      Visibility <- "DB939_Tool_alloc_HMI_Limit_allocation_list"
   Button "Button_96" at 118,470 size 306x41; TextOff 'Text'
      on Press: SetTag("DB939_Tool_alloc_HMI_Selected_prog", 9)
      Visibility <- "DB939_Tool_alloc_HMI_Limit_allocation_list"
   Button "Button_97" at 118,510 size 306x41; TextOff 'Text'
      on Press: SetTag("DB939_Tool_alloc_HMI_Selected_prog", 10)
      Visibility <- "DB939_Tool_alloc_HMI_Limit_allocation_list"
   Button "Button_98" at 118,550 size 306x41; TextOff 'Text'
      on Press: SetTag("DB939_Tool_alloc_HMI_Selected_prog", 11)
      Visibility <- "DB939_Tool_alloc_HMI_Limit_allocation_list"
   Button "Button_99" at 118,590 size 306x41; TextOff 'Text'
      on Press: SetTag("DB939_Tool_alloc_HMI_Selected_prog", 12)
      Visibility <- "DB939_Tool_alloc_HMI_Limit_allocation_list"
   Button "Button_100" at 118,630 size 306x41; TextOff 'Text'
      on Press: SetTag("DB939_Tool_alloc_HMI_Selected_prog", 13)
      Visibility <- "DB939_Tool_alloc_HMI_Limit_allocation_list"
   Button "Button_101" at 118,670 size 306x41; TextOff 'Text'
      on Press: SetTag("DB939_Tool_alloc_HMI_Selected_prog", 14)
      Visibility <- "DB939_Tool_alloc_HMI_Limit_allocation_list"
   Button "Button_102" at 118,710 size 306x41; TextOff 'Text'
      on Press: SetTag("DB939_Tool_alloc_HMI_Selected_prog", 15)
      Visibility <- "DB939_Tool_alloc_HMI_Limit_allocation_list"
   Button "Button_103" at 491,149 size 306x41; TextOff 'Text'
      on Press: SetTag("DB939_Tool_alloc_HMI_Selected_prog", 16)
      Visibility <- "DB939_Tool_alloc_HMI_Limit_allocation_list"
   Button "Button_104" at 491,189 size 306x41; TextOff 'Text'
      on Press: SetTag("DB939_Tool_alloc_HMI_Selected_prog", 17)
      Visibility <- "DB939_Tool_alloc_HMI_Limit_allocation_list"
   Button "Button_105" at 491,229 size 306x41; TextOff 'Text'
      on Press: SetTag("DB939_Tool_alloc_HMI_Selected_prog", 18)
      Visibility <- "DB939_Tool_alloc_HMI_Limit_allocation_list"
   Button "Button_106" at 491,269 size 306x41; TextOff 'Text'
      on Press: SetTag("DB939_Tool_alloc_HMI_Selected_prog", 19)
      Visibility <- "DB939_Tool_alloc_HMI_Limit_allocation_list"
   Button "Button_107" at 491,309 size 306x41; TextOff 'Text'
      on Press: SetTag("DB939_Tool_alloc_HMI_Selected_prog", 20)
      Visibility <- "DB939_Tool_alloc_HMI_Limit_allocation_list"
   Button "Button_108" at 491,349 size 306x41; TextOff 'Text'
      on Press: SetTag("DB939_Tool_alloc_HMI_Selected_prog", 21)
      Visibility <- "DB939_Tool_alloc_HMI_Limit_allocation_list"
   Button "Button_109" at 491,389 size 306x41; TextOff 'Text'
      on Press: SetTag("DB939_Tool_alloc_HMI_Selected_prog", 22)
      Visibility <- "DB939_Tool_alloc_HMI_Limit_allocation_list"
   Button "Button_110" at 491,429 size 306x41; TextOff 'Text'
      on Press: SetTag("DB939_Tool_alloc_HMI_Selected_prog", 23)
      Visibility <- "DB939_Tool_alloc_HMI_Limit_allocation_list"
   Button "Button_111" at 491,469 size 306x41; TextOff 'Text'
      on Press: SetTag("DB939_Tool_alloc_HMI_Selected_prog", 24)
      Visibility <- "DB939_Tool_alloc_HMI_Limit_allocation_list"
   Button "Button_112" at 491,509 size 306x41; TextOff 'Text'
      on Press: SetTag("DB939_Tool_alloc_HMI_Selected_prog", 25)
      Visibility <- "DB939_Tool_alloc_HMI_Limit_allocation_list"
   Button "Button_113" at 491,549 size 306x41; TextOff 'Text'
      on Press: SetTag("DB939_Tool_alloc_HMI_Selected_prog", 26)
      Visibility <- "DB939_Tool_alloc_HMI_Limit_allocation_list"
   Button "Button_114" at 491,589 size 306x41; TextOff 'Text'
      on Press: SetTag("DB939_Tool_alloc_HMI_Selected_prog", 27)
      Visibility <- "DB939_Tool_alloc_HMI_Limit_allocation_list"
   Button "Button_115" at 491,629 size 306x41; TextOff 'Text'
      on Press: SetTag("DB939_Tool_alloc_HMI_Selected_prog", 28)
      Visibility <- "DB939_Tool_alloc_HMI_Limit_allocation_list"
   Button "Button_116" at 491,669 size 306x41; TextOff 'Text'
      on Press: SetTag("DB939_Tool_alloc_HMI_Selected_prog", 29)
      Visibility <- "DB939_Tool_alloc_HMI_Limit_allocation_list"
   Button "Button_117" at 491,709 size 306x41; TextOff 'Text'
      on Press: SetTag("DB939_Tool_alloc_HMI_Selected_prog", 30)
      Visibility <- "DB939_Tool_alloc_HMI_Limit_allocation_list"

screen "0013_Archive Alarm" 1280x800, template "Navigation"
   on GenerateScreen: SetTag("CopyLogControl", 0)
   on ClearScreen: SetTag("NavScreenChange", 0); SetTag("CopyLogControl", 0)
   AlarmView "Alarm Archived Fault" at 108,175 size 1058x498; AlarmLog "Archivanzeige"
      Visibility <- "Archived Alarm Control"
   Button "b_System" at 799,713 size 60x60; TextOff 'System'; PictureOff "system messages"; TextList "ico"; PictureList "ico_System_message"
      Appearance <- "Archived Alarm Control"
      on Click: SetTag("Archived Alarm Control", 3)
      ProcessValue <- "Archived Alarm Control"
   Button "b_Foaming" at 891,712 size 60x60; TextOff 'Foaming'; PictureList "ico_Foaming"
      Appearance <- "Archived Alarm Control"
      on Click: SetTag("Archived Alarm Control", 2)
      ProcessValue <- "Archived Alarm Control"
   Button "b_FaultFoam" at 984,712 size 60x60; TextOff 'Fault/Foam'; PictureList "ico_ActualFault_Foaming"
      Appearance <- "Archived Alarm Control"
      on Click: SetTag("Archived Alarm Control", 1)
      ProcessValue <- "Archived Alarm Control"
   Button "b_Fault" at 1077,712 size 60x60; TextOff 'Fault'; PictureList "ico_Actual_Fault"
      Appearance <- "Archived Alarm Control"
      on Click: SetTag("Archived Alarm Control", 0)
      ProcessValue <- "Archived Alarm Control"
   Button "Button_3" at 326,104 size 451x32; TextOff 'Actual Fault / foaming data'; TextList "Archived_Screen_Name_List"
      ProcessValue <- "Archived Alarm Control"
   Button "b_USB" at 705,712 size 60x60; TextOff 'Export USB'; PictureOff "USB_1"
      on Click: function_e9be9208(1, "Archivanzeige", '\Storage Card USB\', 0)
   Button "b_Fault_1" at 1077,712 size 60x60; TextOff 'Fault'
      on Click: SetTag("Archived Alarm Control", 0)
      Appearance <- "Archived Alarm Control"
   Button "b_Foaming_1" at 891,712 size 60x60; TextOff 'Foaming'
      on Click: SetTag("Archived Alarm Control", 2)
      Appearance <- "Archived Alarm Control"
   Button "b_FaultFoam_1" at 984,712 size 60x60; TextOff 'Fault/Foam'
      on Click: SetTag("Archived Alarm Control", 1)
      Appearance <- "Archived Alarm Control"
   Button "b_System_1" at 799,713 size 60x60; TextOff 'System'; PictureOff "system messages"
      on Click: SetTag("Archived Alarm Control", 3)
      Appearance <- "Archived Alarm Control"
   Button "b_ShifProto_ShotCounter_1" at 208,713 size 60x60; TextOff 'Shot Counter'; PictureList "ico_ShiftProtocol"
      ProcessValue <- "Recipe_Appearance_Control"
      Appearance <- "Recipe_Appearance_Control"
   Button "b_Shiftproto_shiftproto" at 208,713 size 60x60; TextOff 'Shift proto'
      on Click: ActivateScreen("0112_Shift protocol", 0); SetTag("Recipe_Appearance_Control", 2)
      Appearance <- "Recipe_Appearance_Control"
   Button "b_SC" at 478,713 size 60x60; TextOff 'Shot Counter'; PictureList "ico_ShotCounter"
      on Press: ActivateScreen("0891_Shotcounter MixingHead", 0); SetTag("Recipe_Appearance_Control", 5)
      Appearance <- "Recipe_Appearance_Control"
      ProcessValue <- "Recipe_Appearance_Control"
   Button "b_SC_1" at 478,713 size 60x60; TextOff 'Shot Counter'
      on Click: ActivateScreen("0891_Shotcounter MixingHead", 0); SetTag("Recipe_Appearance_Control", 5)
      Appearance <- "Recipe_Appearance_Control"
   Button "b_Shift_Plan" at 118,713 size 60x60; TextOff 'Shift Plan'; PictureList "ico_ShiftPlan"
      on Press: ActivateScreen("0113_SettingShiftPlan", 0); SetTag("Recipe_Appearance_Control", 1)
      Appearance <- "Recipe_Appearance_Control"
      ProcessValue <- "Recipe_Appearance_Control"
   Button "b_Shift_Plan_1" at 118,713 size 60x60; TextOff 'Shift Plan'
      on Click: "SettingShiftPlan"(); ActivateScreen("0113_SettingShiftPlan", 0); SetTag("Recipe_Appearance_Control", 1)
      Appearance <- "Recipe_Appearance_Control"
   Button "b_LS_Lastshot" at 298,713 size 60x60; TextOff 'Last Shot'; PictureList "ico_LastShot"
      on Press: ActivateScreen("0036_Last Shot", 0); SetTag("Recipe_Appearance_Control", 3)
      Appearance <- "Recipe_Appearance_Control"
      ProcessValue <- "Recipe_Appearance_Control"
   Button "b_LS_Lastshot_1" at 298,713 size 60x60; TextOff 'Last Shot'
      on Click: ActivateScreen("0036_Last Shot", 0); SetTag("Recipe_Appearance_Control", 3)
      Appearance <- "Recipe_Appearance_Control"
   Button "b_Consumtion" at 388,713 size 60x60; TextOff 'Consumtion / Consum'; PictureList "ico_consum"
      on Press: ActivateScreen("0890_Consumption", 0); SetTag("Recipe_Appearance_Control", 4)
      Appearance <- "Recipe_Appearance_Control"
      ProcessValue <- "Recipe_Appearance_Control"
   Button "b_Consumtion_1" at 388,713 size 60x60; TextOff 'Consumtion / Consum'
      on Click: ActivateScreen("0890_Consumption", 0); SetTag("Recipe_Appearance_Control", 4)
      Appearance <- "Recipe_Appearance_Control"
   AlarmView "Alarm Archived Fault/Foaming Data" at 108,175 size 1058x498; AlarmLog "Archivanzeige"
      Visibility <- "Archived Alarm Control"
   AlarmView "Alarm Archived Foaming Data" at 108,175 size 1058x498; AlarmLog "Archivanzeige"
      Visibility <- "Archived Alarm Control"
   AlarmView "System Alarm" at 108,175 size 1058x498; AlarmLog "Archivanzeige"
      Visibility <- "Archived Alarm Control"

screen "0006_Tank" 1280x800, template "Navigation"
   on GenerateScreen: SetBit("DB612_Tank_State.Read"); SetTag("Navigation_7", 3)
   Button "Button_6" at 486,558 size 395x220; TextOff 'Text'
      Visibility <- "Tank_Visibility Control"
   TextField "Text field_17" at 576,564 size 184x29; Text 'Tempering tank'
      Visibility <- "Tank_Visibility Control"
   TextField "Text field_18" at 495,600 size 72x25; Text 'Actual:'
      Visibility <- "Tank_Visibility Control"
   TextField "Text field_19" at 493,626 size 100x25; Text 'Set value:'
      Visibility <- "Tank_Visibility Control"
   TextField "Text field_20" at 493,653 size 116x25; Text 'Cooling On:'
      Visibility <- "Tank_Visibility Control"
   TextField "Text field_21" at 493,680 size 120x25; Text 'Cooling Off:'
      Visibility <- "Tank_Visibility Control"
   TextField "Text field_22" at 493,707 size 122x25; Text 'Heating Off:'
      Visibility <- "Tank_Visibility Control"
   TextField "Text field_23" at 493,734 size 118x25; Text 'Heating On:'
      Visibility <- "Tank_Visibility Control"
   IOField "I/O field_11" at 742,600 size 80x25; FormatPattern 999.9
      Visibility <- "Tank_Visibility Control"
      ProcessValue <- "DB602_PV_Tank_Tank{0}_Temp_PV_ActV_Value"
   IOField "I/O field_12" at 742,626 size 80x25; Authorization "Operate"; FormatPattern 999.9
      Visibility <- "Tank_Visibility Control"
      ProcessValue <- "DB602_PV_Tank_Tank{0}_Temp_PV_SetV_Value"
   IOField "I/O field_13" at 742,653 size 80x25; Authorization "Operate"; FormatPattern 999.9
      ProcessValue <- "DB702_Tank_Value.Pt2_Controller[0].Dif_Cooling_ON"
      Visibility <- "Tank_Visibility Control"
   IOField "I/O field_14" at 742,680 size 80x25; Authorization "Operate"; FormatPattern 999.9
      ProcessValue <- "DB702_Tank_Value.Pt2_Controller[0].Dif_Cooling_OFF"
      Visibility <- "Tank_Visibility Control"
   IOField "I/O field_15" at 742,707 size 80x25; Authorization "Operate"; FormatPattern 999.9
      ProcessValue <- "DB702_Tank_Value.Pt2_Controller[0].Dif_Heating_OFF"
      Visibility <- "Tank_Visibility Control"
   IOField "I/O field_16" at 742,734 size 80x25; Authorization "Operate"; FormatPattern 999.9
      ProcessValue <- "DB702_Tank_Value.Pt2_Controller[0].Dif_Heating_ON"
      Visibility <- "Tank_Visibility Control"
   Button "Button_7" at 825,562 size 51x41; TextOff 'Text'; PictureOff "images (1)"
      on Press: SetTag("Tank_Visibility Control", 0)
      Visibility <- "Tank_Visibility Control"
   TextField "Text field_60" at 832,626 size 46x25; Text 'ºC'
      Visibility <- "Tank_Visibility Control"
   TextField "Text field_61" at 832,655 size 41x22; Text 'Δ ºC'
      Visibility <- "Tank_Visibility Control"
   TextField "Text field_62" at 832,600 size 46x25; Text 'ºC'
      Visibility <- "Tank_Visibility Control"
   TextField "Text field_63" at 832,682 size 41x22; Text 'Δ ºC'
      Visibility <- "Tank_Visibility Control"
   TextField "Text field_64" at 832,709 size 41x22; Text 'Δ ºC'
      Visibility <- "Tank_Visibility Control"
   TextField "Text field_65" at 832,736 size 41x22; Text 'Δ ºC'
      Visibility <- "Tank_Visibility Control"
   Button "Button_10" at 486,558 size 395x240; TextOff 'Text'
      Visibility <- "Tank_Visibility Control"
   TextField "Text field_24" at 576,564 size 199x29; Text 'Filling Level tank'
      Visibility <- "Tank_Visibility Control"
   TextField "Text field_25" at 495,598 size 72x25; Text 'Actual:'
      Visibility <- "Tank_Visibility Control"
   TextField "Text field_26" at 495,624 size 99x25; Text 'Max.Level'
      Visibility <- "Tank_Visibility Control"
   TextField "Text field_27" at 495,651 size 114x25; Text 'Stop Filling'
      Visibility <- "Tank_Visibility Control"
   TextField "Text field_28" at 495,678 size 124x25; Text 'Start Filling:'
      Visibility <- "Tank_Visibility Control"
   TextField "Text field_29" at 495,705 size 225x25; Text 'Stop Level stirrer tank:'
      Visibility <- "Tank_Visibility Control"
   TextField "Text field_30" at 495,732 size 187x25; Text 'Warning Min.Level:'
      Visibility <- "Tank_Visibility Control"
   IOField "I/O field_17" at 742,598 size 80x25; FormatPattern 999.9
      Visibility <- "Tank_Visibility Control"
      ProcessValue <- "DB602_PV_Tank_Tank{0}_Level_PV_ActV_Value"
   IOField "I/O field_18" at 742,624 size 80x25; Authorization "Operate"; FormatPattern 999.9
      ProcessValue <- "DB702_Tank_Value.Tank[0].TankLevel.Max_Level"
      Visibility <- "Tank_Visibility Control"
   IOField "I/O field_19" at 742,651 size 80x25; Authorization "Operate"; FormatPattern 999.9
      ProcessValue <- "DB702_Tank_Value.Tank[0].TankLevel.Stop_Level_Filling"
      Visibility <- "Tank_Visibility Control"
   IOField "I/O field_20" at 742,678 size 80x25; Authorization "Operate"; FormatPattern 999.9
      ProcessValue <- "DB702_Tank_Value.Tank[0].TankLevel.Start_Level_Filling"
      Visibility <- "Tank_Visibility Control"
   IOField "I/O field_21" at 742,705 size 80x25; Authorization "Operate"; FormatPattern 999.9
      ProcessValue <- "DB702_Tank_Value.Tank[0].TankLevel.Stop_Level_Agitator"
      Visibility <- "Tank_Visibility Control"
   IOField "I/O field_22" at 742,732 size 80x25; Authorization "Operate"; FormatPattern 999.9
      ProcessValue <- "DB702_Tank_Value.Tank[0].TankLevel.Min_Level_Warning"
      Visibility <- "Tank_Visibility Control"
   Button "Button_11" at 825,562 size 51x41; TextOff 'Text'; PictureOff "images (1)"
      on Press: SetTag("Tank_Visibility Control", 0)
      Visibility <- "Tank_Visibility Control"
   TextField "Text field_31" at 495,758 size 103x25; Text 'Min. level:'
      Visibility <- "Tank_Visibility Control"
   IOField "I/O field_23" at 742,758 size 80x25; Authorization "Operate"; FormatPattern 999.9
      ProcessValue <- "DB702_Tank_Value.Tank[0].TankLevel.Min_Level"
      Visibility <- "Tank_Visibility Control"
   TextField "Text field_33" at 837,598 size 46x25; Text '%'
      Visibility <- "Tank_Visibility Control"
   TextField "Text field_34" at 837,624 size 46x25; Text '%'
      Visibility <- "Tank_Visibility Control"
   TextField "Text field_35" at 837,651 size 46x25; Text '%'
      Visibility <- "Tank_Visibility Control"
   TextField "Text field_36" at 837,678 size 46x25; Text '%'
      Visibility <- "Tank_Visibility Control"
   TextField "Text field_37" at 837,705 size 46x25; Text '%'
      Visibility <- "Tank_Visibility Control"
   TextField "Text field_38" at 837,732 size 46x25; Text '%'
      Visibility <- "Tank_Visibility Control"
   TextField "Text field_39" at 837,758 size 46x25; Text '%'
      Visibility <- "Tank_Visibility Control"
   Button "Template_Button_41" at 16,724 size 68x66; TextOff 'Text'; PictureList "Ico_navigation_2"; PictureOff "Setting_Nav_7"; Authorization "User administration"
      ProcessValue <- "Nav_7"
      on Click: ActivateScreen("0007_Tank Setting", 0)
      Visibility <- "NavUserChange"
   Button "Button_12" at 486,558 size 395x220; TextOff 'Text'
      Visibility <- "Tank_Visibility Control"
   TextField "Text field_45" at 576,564 size 226x29; Text 'Temperature barrel'
      Visibility <- "Tank_Visibility Control"
   TextField "Text field_46" at 495,600 size 72x25; Text 'Actual:'
      Visibility <- "Tank_Visibility Control"
   TextField "Text field_47" at 495,626 size 100x25; Text 'Set value:'
      Visibility <- "Tank_Visibility Control"
   TextField "Text field_49" at 495,680 size 120x25; Text 'Cooling Off:'
      Visibility <- "Tank_Visibility Control"
   TextField "Text field_50" at 495,706 size 122x25; Text 'Heating Off:'
      Visibility <- "Tank_Visibility Control"
   TextField "Text field_51" at 495,733 size 118x25; Text 'Heating On:'
      Visibility <- "Tank_Visibility Control"
   IOField "I/O field_28" at 742,600 size 80x25; FormatPattern 999.9
      Visibility <- "Tank_Visibility Control"
      ProcessValue <- "DB602_PV_Tank_Tank{0}_JacketHeater_PV_ActV_Value"
   IOField "I/O field_29" at 742,626 size 80x25; Authorization "Operate"; FormatPattern 999.9
      Visibility <- "Tank_Visibility Control"
      ProcessValue <- "DB602_PV_Tank_Tank{0}_JacketHeater_PV_SetV_Value"
   IOField "I/O field_31" at 742,680 size 80x25; Authorization "Operate"; FormatPattern 999.9
      Visibility <- "Tank_Visibility Control"
      ProcessValue <- "DB702_Tank_Value_Pt2_ControllerBarell{0}_Dif_Cooling_OFF"
   IOField "I/O field_32" at 742,706 size 80x25; Authorization "Operate"; FormatPattern 999.9
      Visibility <- "Tank_Visibility Control"
      ProcessValue <- "DB702_Tank_Value_Pt2_ControllerBarell{0}_Dif_Heating_OFF"
   IOField "I/O field_33" at 742,733 size 80x25; Authorization "Operate"; FormatPattern 999.9
      Visibility <- "Tank_Visibility Control"
      ProcessValue <- "DB702_Tank_Value_Pt2_ControllerBarell{0}_Dif_Heating_ON"
   Button "Button_13" at 825,562 size 51x41; TextOff 'Text'; PictureOff "images (1)"
      on Press: SetTag("Tank_Visibility Control", 0)
      Visibility <- "Tank_Visibility Control"
   TextField "Text field_54" at 495,653 size 116x25; Text 'Cooling On:'
      Visibility <- "Tank_Visibility Control"
   IOField "I/O field_30" at 742,653 size 80x25; Authorization "Operate"; FormatPattern 999.9
      ProcessValue <- "DB702_Tank_Value_Pt2_ControllerBarell{0}_Dif_Cooling_ON"
      Visibility <- "Tank_Visibility Control"
   TextField "Text field_48" at 832,626 size 46x25; Text 'ºC'
      Visibility <- "Tank_Visibility Control"
   TextField "Text field_52" at 832,655 size 41x22; Text 'Δ ºC'
      Visibility <- "Tank_Visibility Control"
   TextField "Text field_53" at 832,600 size 46x25; Text 'ºC'
      Visibility <- "Tank_Visibility Control"
   TextField "Text field_55" at 832,682 size 41x22; Text 'Δ ºC'
      Visibility <- "Tank_Visibility Control"
   TextField "Text field_56" at 832,708 size 41x22; Text 'Δ ºC'
      Visibility <- "Tank_Visibility Control"
   TextField "Text field_57" at 832,735 size 41x22; Text 'Δ ºC'
      Visibility <- "Tank_Visibility Control"
   Button "Button_3" at 486,558 size 395x220; TextOff 'Text'
      Visibility <- "Tank_Visibility Control"
   TextField "Text field_73" at 576,564 size 210x29; Text 'Temperature tank'
      Visibility <- "Tank_Visibility Control"
   TextField "Text field_74" at 495,600 size 72x25; Text 'Actual:'
      Visibility <- "Tank_Visibility Control"
   TextField "Text field_75" at 495,626 size 100x25; Text 'Set value:'
      Visibility <- "Tank_Visibility Control"
   TextField "Text field_76" at 495,680 size 199x25; Text 'Warning lower limit:'
      Visibility <- "Tank_Visibility Control"
   TextField "Text field_77" at 495,707 size 170x25; Text 'Fault upper limit:'
      Visibility <- "Tank_Visibility Control"
   TextField "Text field_78" at 495,734 size 168x25; Text 'Fault lower limit:'
      Visibility <- "Tank_Visibility Control"
   IOField "I/O field_36" at 742,600 size 80x25; FormatPattern 999.9
      Visibility <- "Tank_Visibility Control"
      ProcessValue <- "DB602_PV_Tank_Tank{0}_Temp_PV_ActV_Value"
   IOField "I/O field_37" at 742,626 size 80x25; Authorization "Operate"; FormatPattern 999.9
      Visibility <- "Tank_Visibility Control"
      ProcessValue <- "DB602_PV_Tank_Tank{0}_Temp_PV_SetV_Value"
   IOField "I/O field_38" at 742,680 size 80x25; Authorization "Operate"; FormatPattern 999.9
      Visibility <- "Tank_Visibility Control"
      ProcessValue <- "DB602_PV_Tank_Tank{0}_Temp_PV_SetV_WarningLowerLimit"
   IOField "I/O field_39" at 742,707 size 80x25; Authorization "Operate"; FormatPattern 999.9
      Visibility <- "Tank_Visibility Control"
      ProcessValue <- "DB602_PV_Tank_Tank{0}_Temp_PV_SetV_AlarmUpperLimit"
   IOField "I/O field_40" at 742,734 size 80x25; Authorization "Operate"; FormatPattern 999.9
      Visibility <- "Tank_Visibility Control"
      ProcessValue <- "DB602_PV_Tank_Tank{0}_Temp_PV_SetV_AlarmLowerLimit"
   Button "Button_21" at 825,562 size 51x41; TextOff 'Text'; PictureOff "images (1)"
      on Press: SetTag("Tank_Visibility Control", 0)
      Visibility <- "Tank_Visibility Control"
   TextField "Text field_80" at 832,626 size 46x25; Text 'ºC'
      Visibility <- "Tank_Visibility Control"
   TextField "Text field_84" at 495,653 size 201x25; Text 'Warning upper limit:'
      Visibility <- "Tank_Visibility Control"
   IOField "I/O field_41" at 742,653 size 80x25; Authorization "Operate"; FormatPattern 999.9
      Visibility <- "Tank_Visibility Control"
      ProcessValue <- "DB602_PV_Tank_Tank{0}_Temp_PV_SetV_WarningUpperLimit"
   TextField "Text field_86" at 832,655 size 41x22; Text 'Δ ºC'
      Visibility <- "Tank_Visibility Control"
   TextField "Text field_79" at 832,600 size 46x25; Text 'ºC'
      Visibility <- "Tank_Visibility Control"
   TextField "Text field_81" at 832,682 size 41x22; Text 'Δ ºC'
      Visibility <- "Tank_Visibility Control"
   TextField "Text field_82" at 832,709 size 41x22; Text 'Δ ºC'
      Visibility <- "Tank_Visibility Control"
   TextField "Text field_83" at 832,736 size 41x22; Text 'Δ ºC'
      Visibility <- "Tank_Visibility Control"
   Button "Button_22" at 486,558 size 395x220; TextOff 'Text'
      Visibility <- "Tank_Visibility Control"
   TextField "Text field_112" at 576,564 size 202x29; Text 'Nucleation tank:'
      Visibility <- "Tank_Visibility Control"
   TextField "Text field_113" at 495,600 size 72x25; Text 'Actual:'
      Visibility <- "Tank_Visibility Control"
   TextField "Text field_114" at 495,626 size 100x25; Text 'Set value:'
      Visibility <- "Tank_Visibility Control"
   TextField "Text field_115" at 495,680 size 199x25; Text 'Warning lower limit:'
      Visibility <- "Tank_Visibility Control"
   TextField "Text field_116" at 495,706 size 170x25; Text 'Fault upper limit:'
      Visibility <- "Tank_Visibility Control"
   TextField "Text field_117" at 495,733 size 168x25; Text 'Fault lower limit:'
      Visibility <- "Tank_Visibility Control"
   IOField "I/O field_42" at 742,600 size 80x25; FormatPattern 999.9
      Visibility <- "Tank_Visibility Control"
      ProcessValue <- "DB602_PV_Tank_Tank{0}_Nucleation_PV_ActV_Value"
   IOField "I/O field_44" at 742,626 size 80x25; Authorization "Operate"; FormatPattern 999.9
      Visibility <- "Tank_Visibility Control"
      ProcessValue <- "DB602_PV_Tank_Tank{0}_Nucleation_PV_SetV_Value"
   IOField "I/O field_45" at 742,680 size 80x25; Authorization "Operate"; FormatPattern 999.9
      Visibility <- "Tank_Visibility Control"
      ProcessValue <- "DB602_PV_Tank_Tank{0}_Nucleation_PV_SetV_WarningLowerLimit"
   IOField "I/O field_46" at 742,706 size 80x25; Authorization "Operate"; FormatPattern 999.9
      Visibility <- "Tank_Visibility Control"
      ProcessValue <- "DB602_PV_Tank_Tank{0}_Nucleation_PV_SetV_AlarmLowerLimit"
   IOField "I/O field_47" at 742,733 size 80x25; Authorization "Operate"; FormatPattern 999.9
      Visibility <- "Tank_Visibility Control"
      ProcessValue <- "DB602_PV_Tank_Tank{0}_Nucleation_PV_SetV_AlarmUpperLimit"
   Button "Button_23" at 825,562 size 51x41; TextOff 'Text'; PictureOff "images (1)"
      on Press: SetTag("Tank_Visibility Control", 0)
      Visibility <- "Tank_Visibility Control"
   TextField "Text field_118" at 832,600 size 46x25; Text '%'
      Visibility <- "Tank_Visibility Control"
   TextField "Text field_119" at 832,626 size 46x25; Text '%'
      Visibility <- "Tank_Visibility Control"
   TextField "Text field_123" at 495,653 size 201x25; Text 'Warning upper limit:'
      Visibility <- "Tank_Visibility Control"
   IOField "I/O field_48" at 742,653 size 80x25; Authorization "Operate"; FormatPattern 999.9
      Visibility <- "Tank_Visibility Control"
      ProcessValue <- "DB602_PV_Tank_Tank{0}_Nucleation_PV_SetV_WarningUpperLimit"
   TextField "Text field_125" at 832,655 size 40x22; Text 'Δ %'
      Visibility <- "Tank_Visibility Control"
   TextField "Text field_71" at 832,682 size 40x22; Text 'Δ %'
      Visibility <- "Tank_Visibility Control"
   TextField "Text field_72" at 832,708 size 40x22; Text 'Δ %'
      Visibility <- "Tank_Visibility Control"
   TextField "Text field_120" at 832,735 size 40x22; Text 'Δ %'
      Visibility <- "Tank_Visibility Control"
   Button "b_Tank2" at 160,608 size 48x32; TextOff 'Text'
      on Press: ActivateScreen("0024_ActualFaults", 0); SetTag("Alarm_Filter_Tag", 4); SetTag("NavScreenChange", 0)
      ObjectEnable <- "DB612_Tank_State_FaultExists{2}"
   Button "b_Tank2_1" at 155,351 size 48x32; TextOff 'Text'
      on Press: ActivateScreen("0024_ActualFaults", 0); SetTag("Alarm_Filter_Tag", 4)
      ObjectEnable <- "DB612_Tank_State_FaultExists{2}"
   Button "b_Tank1" at 248,480 size 39x32; TextOff 'Text'
      on Press: ActivateScreen("0024_ActualFaults", 0); SetTag("Alarm_Filter_Tag", 4); SetTag("NavScreenChange", 0)
      ObjectEnable <- "DB612_Tank_State_FaultExists{1}"
   TextField "Text field_58" at 316,210 size 89x25; Text '°C'
      Visibility <- "DB702_Tank_Value_Tank{0}_With_BarelStation_Heating"
   TextField "Text field_14" at 363,474 size 80x25; Text '°C'
   TextField "Text field_70" at 363,534 size 80x25; Text '%'
      Visibility <- "DB702_Tank_Value_Tank{0}_With_Nucleation"
   Button "Button_1" at 485,151 size 395x401; TextOff 'Text'
   TextField "Text field_1" at 493,164 size 77x25; Text 'Density'
   TextField "Text field_2" at 493,187 size 204x25; Text 'Runtime stirrer tank:'
      Visibility <- "DB702_Tank_Value_Tank{0}_With_Agitator"
   TextField "Text field_3" at 493,213 size 227x25; Text 'Break time stirrer tank:'
      Visibility <- "DB702_Tank_Value_Tank{0}_With_Agitator"
   TextField "Text field_4" at 493,265 size 166x25; Text 'Max. filling time:'
      Visibility <- "DB702_Tank_Value_Tank{0}_With_Filling"
   TextField "Text field_5" at 493,291 size 171x25; Text 'Filling after shot:'
      Visibility <- "DB702_Tank_Value_Tank{0}_With_Filling"
   TextField "Text field_6" at 493,317 size 171x25; Text 'Filling after time:'
      Visibility <- "DB702_Tank_Value_Tank{0}_With_Filling"
   TextField "Text field_7" at 493,343 size 212x25; Text 'set temperature tank:'
   IOField "Tank_IO_Density" at 712,161 size 90x25; Authorization "User administration"; FormatPattern 9999
      ProcessValue <- "DB702_Tank_Value.Tank[0].Density"
   IOField "I/O field_2" at 722,187 size 80x25; Authorization "Operate"; FormatPattern 99999
      ProcessValue <- "DB702_Tank_Value_Tank{0}_Agitator_RunTime"
      Visibility <- "DB702_Tank_Value_Tank{0}_With_Agitator"
   IOField "I/O field_3" at 722,213 size 80x25; Authorization "Operate"; FormatPattern 99999
      ProcessValue <- "DB702_Tank_Value_Tank{0}_Agitator_PauseTime"
      Visibility <- "DB702_Tank_Value_Tank{0}_With_Agitator"
   IOField "I/O field_4" at 722,265 size 80x25; Authorization "Operate"; FormatPattern 99999
      ProcessValue <- "DB702_Tank_Value_Tank{0}_FillingTimeControl"
      Visibility <- "DB702_Tank_Value_Tank{0}_With_Filling"
   IOField "I/O field_5" at 722,291 size 80x25; Authorization "Operate"; FormatPattern 999
      ProcessValue <- "DB702_Tank_Value_Tank{0}_NoShotFilling"
      Visibility <- "DB702_Tank_Value_Tank{0}_With_Filling"
   IOField "I/O field_6" at 722,317 size 80x25; Authorization "Operate"; FormatPattern 99999
      ProcessValue <- "DB702_Tank_Value_Tank{0}_TimeToStartFilling"
      Visibility <- "DB702_Tank_Value_Tank{0}_With_Filling"
   IOField "I/O field_7" at 722,343 size 80x25; Authorization "Operate"; FormatPattern 999.9
      ProcessValue <- "DB602_PV_Tank_Tank{0}_Temp_PV_SetV_Value"
   TextField "Text field_8" at 806,161 size 65x25; Text 'g/cm³'
   TextField "Text field_9" at 806,187 size 46x25; Text 's'
      Visibility <- "DB702_Tank_Value_Tank{0}_With_Agitator"
   TextField "Text field_10" at 806,213 size 46x25; Text 's'
      Visibility <- "DB702_Tank_Value_Tank{0}_With_Agitator"
   TextField "Text field_11" at 806,265 size 46x25; Text 's'
      Visibility <- "DB702_Tank_Value_Tank{0}_With_Filling"
   TextField "Text field_12" at 806,317 size 46x25; Text 's'
      Visibility <- "DB702_Tank_Value_Tank{0}_With_Filling"
   TextField "Text field_13" at 806,343 size 46x25; Text 'ºC'
   IOField "I/O field_8" at 363,474 size 56x25; FormatPattern 999.9
      ProcessValue <- "DB602_PV_Tank_Tank{0}_Temp_PV_ActV_Value"
   Button "b_Incress_Tank" at 789,104 size 46x32; TextOff 'Text'; PictureOff "right arrow"
      on Click: function_dd21b452("DB612_Tank_State.ReadDeviceNo", 1)
   Button "b_Decress_Tank" at 269,104 size 46x32; TextOff 'Text'; PictureOff "left arrow"
      on Click: function_b9b71300("DB612_Tank_State.ReadDeviceNo", 1)
   TextField "Text field_15" at 493,369 size 161x25; Text 'Level niveau up:'
      Visibility <- "DB702_Tank_Value_Tank{0}_With_Level_Probe"
   TextField "Text field_16" at 493,395 size 189x25; Text 'Level niveau down:'
      Visibility <- "DB702_Tank_Value_Tank{0}_With_Level_Probe"
   IOField "I/O field_9" at 722,369 size 80x25; Authorization "Operate"; FormatPattern 999.9
      ProcessValue <- "DB702_Tank_Value.Tank[0].TankLevel.Stop_Level_Filling"
      Visibility <- "DB702_Tank_Value_Tank{0}_With_Level_Probe"
   IOField "I/O field_10" at 722,395 size 80x25; Authorization "Operate"; FormatPattern 999.9
      ProcessValue <- "DB702_Tank_Value.Tank[0].TankLevel.Start_Level_Filling"
      Visibility <- "DB702_Tank_Value_Tank{0}_With_Level_Probe"
   Button "b_Tank_SetTemperatureTank" at 830,341 size 45x30; TextOff 'Text'; PictureOff "obeng"
      on Press: SetTag("Tank_Visibility Control", 1)
   Button "b_Tank_Set_Niveau_Up" at 830,367 size 45x30; TextOff 'Text'; PictureOff "obeng"
      on Press: SetTag("Tank_Visibility Control", 2)
      Visibility <- "DB702_Tank_Value_Tank{0}_With_Level_Probe"
   TextField "Text field_32" at 363,504 size 80x25; Text '%'
      Visibility <- "DB702_Tank_Value_Tank{0}_With_Level_Probe"
   TextField "Text field_40" at 806,369 size 46x25; Text '%'
      Visibility <- "DB702_Tank_Value_Tank{0}_With_Level_Probe"
   TextField "Text field_41" at 806,395 size 46x25; Text '%'
      Visibility <- "DB702_Tank_Value_Tank{0}_With_Level_Probe"
   IOField "I/O field_25" at 722,466 size 80x25; Authorization "Operate"; FormatPattern 999.9
      ProcessValue <- "DB602_PV_Tank_Tank{0}_JacketHeater_PV_SetV_Value"
      Visibility <- "DB702_Tank_Value_Tank{0}_With_BarelStation_Heating"
   IOField "I/O field_26" at 722,492 size 80x25; Authorization "Operate"; FormatPattern 99999
      ProcessValue <- "DB702_Tank_Value_CirculationPump{0}_RunTime"
      Visibility <- "DB702_Tank_Value_Tank{0}_With_BarelStation_Zirkulation"
   IOField "I/O field_27" at 722,518 size 80x25; Authorization "Operate"; FormatPattern 99999
      ProcessValue <- "DB702_Tank_Value_CirculationPump{0}_PauseTime"
      Visibility <- "DB702_Tank_Value_Tank{0}_With_BarelStation_Zirkulation"
   TextField "Text field_42" at 493,466 size 228x25; Text 'Set temperature barrel:'
      Visibility <- "DB702_Tank_Value_Tank{0}_With_BarelStation_Heating"
   TextField "Text field_43" at 493,492 size 212x25; Text 'Runtime pump barrel:'
      Visibility <- "DB702_Tank_Value_Tank{0}_With_BarelStation_Zirkulation"
   TextField "Text field_44" at 493,518 size 237x25; Text 'Pause time pump barrel:'
      Visibility <- "DB702_Tank_Value_Tank{0}_With_BarelStation_Zirkulation"
   Button "b_Tank_SetTemperatureBarrel" at 830,464 size 45x30; TextOff 'Text'; PictureOff "obeng"
      on Press: SetTag("Tank_Visibility Control", 3)
      Visibility <- "DB702_Tank_Value_Tank{0}_With_BarelStation_Heating"
   IOField "I/O field_34" at 316,210 size 62x25; FormatPattern 999.9
      ProcessValue <- "DB602_PV_Tank_Tank{0}_JacketHeater_PV_ActV_Value"
      Visibility <- "DB702_Tank_Value_Tank{0}_With_BarelStation_Heating"
   IOField "I/O field_43" at 326,104 size 451x32; Authorization "Operate"; FormatPattern ????????????????????
      ProcessValue <- "DB702_Tank_Value_Tank{0}_Name"
      Appearance <- "DB702_Tank_Value_Tank{0}_Color"
   IOField "I/O field_35" at 363,534 size 56x25; FormatPattern 999.9
      ProcessValue <- "DB602_PV_Tank_Tank{0}_Nucleation_PV_ActV_Value"
      Visibility <- "DB702_Tank_Value_Tank{0}_With_Nucleation"
   Button "Button_24" at 363,474 size 80x25; TextOff 'Text'
      on Press: SetTag("Tank_Visibility Control", 4)
   Button "Button_25" at 363,534 size 80x25; TextOff 'Text'
      on Press: SetTag("Tank_Visibility Control", 5)
      Visibility <- "DB702_Tank_Value_Tank{0}_With_Nucleation"
   IOField "I/O field_49" at 722,239 size 80x25; Authorization "Operate"; FormatPattern 99999
      Visibility <- "DB702_Tank_Value_Tank{0}_With_BarelStation_Zirkulation"
      ProcessValue <- "DB702_Tank_Value_Tank{0}_PreAgitatingTime"
   TextField "Text field_152" at 493,239 size 156x25; Text 'Pre Mixing Time'
      Visibility <- "DB702_Tank_Value_Tank{0}_With_BarelStation_Zirkulation"
   Button "Button_8" at 1081,188 size 81x116; TextOff 'Text'
      Visibility <- "DB702_Tank_Value_Tank{0}_With_Agitator"
   GraphicView "Graphic view_7" at 1093,252 size 56x48; Picture "Agitator"
      Visibility <- "DB702_Tank_Value_Tank{0}_With_Agitator"
   Rectangle "Rectangle_8" at 1090,196 size 64x56
      Appearance <- "DB612_Tank_State_Agitator{0}_State_Drive"
      Visibility <- "DB702_Tank_Value_Tank{0}_With_Agitator"
   GraphicIOField "Graphic I/O field_7" at 1098,199 size 48x48; PictureList "ON_OFF_SWITCH"
      ProcessValue <- "DB612_Tank_State_Agitator{0}_Switch_Drive_ON_OFF"
      Visibility <- "DB702_Tank_Value_Tank{0}_With_Agitator"
   Button "Button_9" at 1079,180 size 88x128; TextOff 'Text'
      on Click: InvertBit("DB612_Tank_State_Agitator{0}_Switch_Drive_ON_OFF")
      Visibility <- "DB702_Tank_Value_Tank{0}_With_Agitator"
   Button "Button_5" at 995,188 size 81x116; TextOff 'Text'
      Visibility <- "DB702_Tank_Value_Tank{0}_With_Filling"
   GraphicView "Graphic view_6" at 1007,252 size 56x48; Picture "Refilling"
      Visibility <- "DB702_Tank_Value_Tank{0}_With_Filling"
   Rectangle "Rectangle_7" at 1003,196 size 64x56
      Appearance <- "DB612_Tank_State_Tank{0}_State_Refilling"
      Visibility <- "DB702_Tank_Value_Tank{0}_With_Filling"
   GraphicIOField "Graphic I/O field_6" at 1011,199 size 48x48; PictureList "ON_OFF_SWITCH"
      ProcessValue <- "DB612_Tank_State_Tank{0}_Switch_Refilling_ON_OFF"
      Visibility <- "DB702_Tank_Value_Tank{0}_With_Filling"
   Button "Button_15" at 992,180 size 88x128; TextOff 'Text'
      on Click: InvertBit("DB612_Tank_State_Tank{0}_Switch_Refilling_ON_OFF")
      Visibility <- "DB702_Tank_Value_Tank{0}_With_Filling"
   Button "Button_4" at 905,187 size 81x116; TextOff 'Text'
   GraphicView "Graphic view_5" at 917,252 size 56x48; Picture "Switch Temp"
   Rectangle "Rectangle_6" at 914,195 size 64x56
      Appearance <- "DB612_Tank_State_ControllerTankTemp{0}_State_Temp"
   GraphicIOField "Graphic I/O field_5" at 922,198 size 48x48; PictureList "ON_OFF_SWITCH"
      ProcessValue <- "DB612_Tank_State_ControllerTankTemp{0}_Switch_Temp_ON_OFF"
   Button "Button_20" at 901,179 size 88x128; TextOff 'Text'
      on Click: InvertBit("DB612_Tank_State_ControllerTankTemp{0}_Switch_Temp_ON_OFF")
   Button "Button_2" at 905,472 size 81x116; TextOff 'Text'
      Visibility <- "DB702_Tank_Value_Tank{0}_With_Filling_2Valve"
   GraphicView "Graphic view_2" at 917,536 size 56x48; Picture "FillingFromBarel"
      Visibility <- "DB702_Tank_Value_Tank{0}_With_Filling_2Valve"
   Rectangle "Rectangle_1" at 913,480 size 64x56
      Visibility <- "DB702_Tank_Value_Tank{0}_With_Filling_2Valve"
      Appearance <- "DB612_Tank_State_Tank{0}_Switch_Refilling_from_Barrel_ON_OFF"
   GraphicIOField "Graphic I/O field_1" at 921,483 size 48x48; PictureList "ON_OFF_SWITCH"
      ProcessValue <- "DB612_Tank_State_Tank{0}_Switch_Refilling_from_Barrel_ON_OFF"
      Visibility <- "DB702_Tank_Value_Tank{0}_With_Filling_2Valve"
   Button "Button_26" at 902,467 size 88x128; TextOff 'Text'
      on Click: InvertBit("DB612_Tank_State_Tank{0}_Switch_Refilling_from_Barrel_ON_OFF")
      Visibility <- "DB702_Tank_Value_Tank{0}_With_Filling_2Valve"
   Button "Button_19" at 906,331 size 81x116; TextOff 'Text'
      Visibility <- "DB702_Tank_Value_Tank{0}_With_BarelStation_Heating"
   GraphicView "Graphic view_3" at 918,396 size 56x48; Picture "HeaJacket"
      Visibility <- "DB702_Tank_Value_Tank{0}_With_BarelStation_Heating"
   Rectangle "Rectangle_3" at 915,339 size 64x56
      Appearance <- "DB612_Tank_State_ControllerBarellTemp{0}_State_Temp"
      Visibility <- "DB702_Tank_Value_Tank{0}_With_BarelStation_Heating"
   GraphicIOField "Graphic I/O field_2" at 923,342 size 48x48; PictureList "ON_OFF_SWITCH"
      ProcessValue <- "DB612_Tank_State_ControllerBarellTemp{0}_Switch_Temp_ON_OFF"
      Visibility <- "DB702_Tank_Value_Tank{0}_With_BarelStation_Heating"
   Button "Button_27" at 902,323 size 88x128; TextOff 'Text'
      on Click: InvertBit("DB612_Tank_State_ControllerBarellTemp{0}_Switch_Temp_ON_OFF")
      Visibility <- "DB702_Tank_Value_Tank{0}_With_BarelStation_Heating"
   Button "Button_16" at 996,472 size 81x116; TextOff 'Text'
      Visibility <- "DB702_Tank_Value_Tank{0}_With_BarelStation_Zirkulation"
   GraphicView "Graphic view_4" at 1008,544 size 56x34; Picture "motor2"
      Visibility <- "DB702_Tank_Value_Tank{0}_With_BarelStation_Zirkulation"
   Rectangle "Rectangle_4" at 1005,480 size 64x56
      Appearance <- "DB612_Tank_State_CirculationPump{0}_State_Drive"
      Visibility <- "DB702_Tank_Value_Tank{0}_With_BarelStation_Zirkulation"
   GraphicIOField "Graphic I/O field_3" at 1013,483 size 48x48; PictureList "ON_OFF_SWITCH"
      ProcessValue <- "DB612_Tank_State_CirculationPump{0}_Switch_Drive_ON_OFF"
      Visibility <- "DB702_Tank_Value_Tank{0}_With_BarelStation_Zirkulation"
   Button "Button_28" at 992,468 size 88x128; TextOff 'Text'
      on Click: InvertBit("DB612_Tank_State_CirculationPump{0}_Switch_Drive_ON_OFF")
      Visibility <- "DB702_Tank_Value_Tank{0}_With_BarelStation_Zirkulation"
   Button "Button_29" at 1081,330 size 81x116; TextOff 'Text'
      Visibility <- "DB702_Tank_Value_Tank{0}_With_Vacuum"
   GraphicView "Graphic view_8" at 1099,395 size 48x48; Picture "Vacum"
      Visibility <- "DB702_Tank_Value_Tank{0}_With_Vacuum"
   Rectangle "Rectangle_5" at 1090,338 size 64x56
      Visibility <- "DB702_Tank_Value_Tank{0}_With_Vacuum"
      Appearance <- "DB612_Tank_State_Vacuum{0}_Status_Vacuum"
   GraphicIOField "Graphic I/O field_4" at 1098,341 size 48x48; PictureList "ON_OFF_SWITCH"
      Visibility <- "DB702_Tank_Value_Tank{0}_With_Vacuum"
      ProcessValue <- "DB612_Tank_State_Vacuum{0}_Switch_Vacuum_ON_OFF"
   Button "Button_30" at 1077,322 size 88x128; TextOff 'Text'
      on Click: InvertBit("DB612_Tank_State_Vacuum{0}_Switch_Vacuum_ON_OFF")
      Visibility <- "DB702_Tank_Value_Tank{0}_With_Vacuum"
   Button "Button_14" at 1084,472 size 81x116; TextOff 'Text'
      Visibility <- "DB702_Tank_Value_Tank{0}_With_Drain"
   GraphicView "Graphic view_9" at 1098,534 size 56x48; Picture "Drain"
      Visibility <- "DB702_Tank_Value_Tank{0}_With_Drain"
   Rectangle "Rectangle_9" at 1093,480 size 64x56
      Appearance <- "DB612_Tank_State_Tank{0}_Switch_DrainTank_ON_OFF"
      Visibility <- "DB702_Tank_Value_Tank{0}_With_Drain"
   GraphicIOField "Graphic I/O field_8" at 1101,483 size 48x48; PictureList "ON_OFF_SWITCH"
      ProcessValue <- "DB612_Tank_State_Tank{0}_Switch_DrainTank_ON_OFF"
      Visibility <- "DB702_Tank_Value_Tank{0}_With_Drain"
   Button "Button_31" at 1080,468 size 88x128; TextOff 'Text'
      on Click: InvertBit("DB612_Tank_State_Tank{0}_Switch_DrainTank_ON_OFF")
      Visibility <- "DB702_Tank_Value_Tank{0}_With_Drain"
   GraphicView "Graphic view_1" at 168,372 size 129x217; Picture "tank"
   GraphicIOField "Graphic I/O field_9" at 188,426 size 20x20; PictureList "Tank_Sensor"
      Visibility <- "DB702_Tank_Value_Tank{0}_With_Level_3Liq"
      ProcessValue <- "DB612_Tank_State_Tank{0}_Stop_Level_Filling"
   GraphicIOField "Graphic I/O field_10" at 188,458 size 20x20; PictureList "Tank_Sensor"
      Visibility <- "DB702_Tank_Value_Tank{0}_With_Level_4Liq"
      ProcessValue <- "DB612_Tank_State_Tank{0}_Start_Level_Filling"
   GraphicIOField "Graphic I/O field_11" at 188,521 size 20x20; PictureList "Tank_Sensor"
      Visibility <- "DB702_Tank_Value_Tank{0}_With_Level_SMin"
      ProcessValue <- "DB612_Tank_State_Tank{0}_Min_Level"
   GraphicIOField "Graphic I/O field_12" at 256,404 size 20x20; PictureList "Tank_Sensor"
      Visibility <- "DB702_Tank_Value_Tank{0}_With_Level_SMax"
      ProcessValue <- "DB612_Tank_State_Tank{0}_Max_Level"
   GraphicIOField "Graphic I/O field_13" at 300,465 size 20x20; PictureList "Tank_Sensor"
      Visibility <- "DB702_Tank_Value_Tank{0}_With_Filling_Switch"
      ProcessValue <- "DB612_Tank_State_Tank{0}_Max_Level"
   GraphicView "Graphic view_10" at 296,404 size 32x45; Picture "Graphic_7"
      Visibility <- "DB702_Tank_Value_Tank{0}_With_Filling_Valve"
   GraphicView "Graphic view_11" at 344,404 size 32x45; Picture "Graphic_7"
      Visibility <- "DB702_Tank_Value_Tank{0}_With_Filling_2Valve"
   GraphicIOField "Graphic I/O field_14" at 344,372 size 25x20; PictureList "Tank_Sensor"
      Visibility <- "DB702_Tank_Value_Tank{0}_With_Filling_Switch"
      ProcessValue <- "DB612_Tank_State_Tank{0}_Max_Level"
   GraphicView "Graphic view_12" at 296,508 size 32x45; Picture "Graphic_7"
      Visibility <- "DB702_Tank_Value_Tank{0}_With_Filling_ShutDown"
   Rectangle "Rectangle_11" at 339,362 size 40x40
      Visibility <- "DB702_Tank_Value_Tank{0}_With_Filling_2Valve"
   GraphicView "Graphic view_15" at 104,468 size 72x117; Picture "HeaterBackFL"
      Visibility <- "DB702_Tank_Value_Tank{0}_With_Tempering_WTRL"
   GraphicView "Graphic view_17" at 256,192 size 75x86; Picture "Graphic_16"
      Visibility <- "DB702_Tank_Value_Tank{0}_With_BarelStation"
   GraphicView "Graphic view_18" at 203,336 size 53x54; Picture "Graphic_17"
      Visibility <- "DB702_Tank_Value_Tank{0}_With_Agitator"
   GraphicView "Graphic view_19" at 120,339 size 26x38; Picture "Graphic_18"
      Visibility <- "DB702_Tank_Value_Tank{0}_With_Agitator_Converter"
   GraphicView "Graphic view_20" at 213,576 size 42x37; Picture "HEATER"
      Visibility <- "DB702_Tank_Value_Tank{0}_With_Tempering_Heizung"
   GraphicView "Graphic view_14" at 120,224 size 104x48; Picture "motor2"
      Visibility <- "DB702_Tank_Value_Tank{0}_With_BarelStation_Zirkulation"
   GraphicView "Graphic view_16" at 288,580 size 82x86; Picture "Graphic_19"
      Visibility <- "DB702_Tank_Value_Tank{0}_With_Tempering_TempGeraet"
   GraphicView "Alarm Indicator Tank1" at 252,480 size 27x26; Picture "AlarmState2"
      Visibility <- "DB612_Tank_State_FaultExists{1}"
   GraphicView "Alarm Indicator Tank2" at 167,608 size 28x25; Picture "AlarmState2"
      Visibility <- "DB612_Tank_State_FaultExists{2}"
   GraphicIOField "Graphic I/O field_15" at 139,397 size 34x30; PictureList "Valve_Tank"
      ProcessValue <- "Internal_Tank_"
      Visibility <- "DB702_Tank_Value_Tank{0}_With_Tempering_VKaltwasser"
   GraphicIOField "Graphic I/O field_16" at 103,560 size 34x30; PictureList "Valve_Tank"
      Visibility <- "DB702_Tank_Value_Tank{0}_With_Tempering_WTRL"
      ProcessValue <- "Internal_Tank_"
   GraphicView "Graphic view_13" at 295,368 size 35x29; Picture "startfilling"
      Visibility <- "DB612_Tank_State_Tank{0}_Filling_Start"
   TextField "Text field_59" at 806,466 size 46x25; Text 'ºC'
      Visibility <- "DB702_Tank_Value_Tank{0}_With_BarelStation_Heating"
   TextField "Text field_85" at 806,492 size 46x25; Text 's'
      Visibility <- "DB702_Tank_Value_Tank{0}_With_BarelStation_Zirkulation"
   TextField "Text field_87" at 806,518 size 46x25; Text 's'
      Visibility <- "DB702_Tank_Value_Tank{0}_With_BarelStation_Zirkulation"
   GraphicIOField "Graphic I/O field_17" at 188,426 size 20x20; PictureList "Tank_Sensor"
      ProcessValue <- "DB612_Tank_State_Tank{0}_Stop_Level_Filling"
      Visibility <- "DB702_Tank_Value_Tank{0}_With_Level_4Liq"
   TextField "Text field_66" at 806,239 size 46x25; Text 's'
      Visibility <- "DB702_Tank_Value_Tank{0}_With_BarelStation_Zirkulation"
   GraphicView "Alarm Indicator Tank2_1" at 162,351 size 28x25; Picture "AlarmState2"
      Visibility <- "DB612_Tank_State_Agitator{0}_FLT_Exist"
   GraphicView "Graphic view_21" at 167,312 size 35x29; Picture "startfilling"
      Visibility <- "DB612_Tank_State_Agitator{0}_Run"
   IOField "I/O field_24" at 363,504 size 56x25; FormatPattern 999.9
      ProcessValue <- "DB602_PV_Tank_Tank{0}_Level_PV_ActV_Value"
      Visibility <- "DB702_Tank_Value_Tank{0}_With_Level_Probe"
   TextField "Text field_67" at 721,434 size 96x22; Text '-------------'
   GraphicView "Graphic view_22" at 296,404 size 32x45; Picture "Graphic_7"
      Visibility <- "DB702_Tank_Value_Tank{0}_With_Filling_ShutDown"
   Rectangle "Rectangle_14" at 219,410 size 33x142
      Visibility <- "DB612_Tank_State_Tank{0}_Max_Level"
   Rectangle "Rectangle_10" at 219,505 size 33x46
      Visibility <- "DB612_Tank_State_Tank{0}_Min_Level"
   Rectangle "Rectangle_13" at 219,429 size 33x122
      Visibility <- "DB612_Tank_State_Tank{0}_Start_Level_Filling"
   Rectangle "Rectangle_12" at 219,409 size 33x142
      Visibility <- "DB612_Tank_State_Tank{0}_Max_Level"
   Bar "Bar_2" at 218,408 size 35x145; MinimumValue 0; MaximumValue 100
      ProcessValue <- "DB602_PV_Tank_Tank{0}_Level_PV_ActV_Value"
      Visibility <- "DB702_Tank_Value_Tank{0}_With_Level_Probe"

